discrete alarms
   1: 'Rockwell PLC Comm Fault', class No Acknowledgement, trigger "DB302_HMI_Faults_SDC_Faults_0" bit 0
   2: 'Wireless Access Point 1 Comm Fault', class No Acknowledgement, trigger "DB302_HMI_Faults_SDC_Faults_0" bit 1
   3: 'Wireless Access Point 2 Comm Fault', class No Acknowledgement, trigger "DB302_HMI_Faults_SDC_Faults_0" bit 2
   5: 'Wireless Access Point 4 Comm Fault', class No Acknowledgement, trigger "DB302_HMI_Faults_SDC_Faults_0" bit 4
   6: 'Wireless Access Point 5 Comm Fault', class No Acknowledgement, trigger "DB302_HMI_Faults_SDC_Faults_0" bit 5
   7: 'Wireless Access Point 6 Comm Fault', class No Acknowledgement, trigger "DB302_HMI_Faults_SDC_Faults_0" bit 6
   8: 'Wireless Access Point 7 Comm Fault', class No Acknowledgement, trigger "DB302_HMI_Faults_SDC_Faults_0" bit 7
   9: 'Wireless Access Point 8 Comm Fault', class No Acknowledgement, trigger "DB302_HMI_Faults_SDC_Faults_0" bit 8
   10: 'Wireless Access Point 9 Comm Fault', class No Acknowledgement, trigger "DB302_HMI_Faults_SDC_Faults_0" bit 9
   11: 'Wireless Access Point 10 Comm Fault', class No Acknowledgement, trigger "DB302_HMI_Faults_SDC_Faults_0" bit 10
   12: 'Wireless Access Point 11 Comm Fault', class No Acknowledgement, trigger "DB302_HMI_Faults_SDC_Faults_0" bit 11
   13: 'Wireless Access Point 12 Comm Fault', class No Acknowledgement, trigger "DB302_HMI_Faults_SDC_Faults_0" bit 12
   14: 'Wireless Access Point 13 Comm Fault', class No Acknowledgement, trigger "DB302_HMI_Faults_SDC_Faults_0" bit 13
   15: 'Wireless Access Point 14 Comm Fault', class No Acknowledgement, trigger "DB302_HMI_Faults_SDC_Faults_0" bit 14
   16: 'Wireless Access Point 15 Comm Fault', class No Acknowledgement, trigger "DB302_HMI_Faults_SDC_Faults_0" bit 15
   17: 'Wireless Access Point 16 Comm Fault', class No Acknowledgement, trigger "DB302_HMI_Faults_SDC_Faults_1" bit 0
   18: 'Wireless Access Point 17 Comm Fault', class No Acknowledgement, trigger "DB302_HMI_Faults_SDC_Faults_1" bit 1
   19: 'Wireless Access Point 18 Comm Fault', class No Acknowledgement, trigger "DB302_HMI_Faults_SDC_Faults_1" bit 2
   20: 'Wireless Access Point 19 Comm Fault', class No Acknowledgement, trigger "DB302_HMI_Faults_SDC_Faults_1" bit 3
   21: 'Spare_Fault_021', class No Acknowledgement, trigger "DB302_HMI_Faults_SDC_Faults_1" bit 4
   22: 'Spare_Fault_022', class No Acknowledgement, trigger "DB302_HMI_Faults_SDC_Faults_1" bit 5
   23: 'Spare_Fault_023', class No Acknowledgement, trigger "DB302_HMI_Faults_SDC_Faults_1" bit 6
   24: 'Spare_Fault_024', class No Acknowledgement, trigger "DB302_HMI_Faults_SDC_Faults_1" bit 7
   25: 'Duplicate Carrier Fault', class No Acknowledgement, trigger "DB302_HMI_Faults_SDC_Faults_1" bit 8
   26: 'Spare_Fault_026', class No Acknowledgement, trigger "DB302_HMI_Faults_SDC_Faults_1" bit 9
   27: 'EMS01 System E-Stop', class No Acknowledgement, trigger "DB302_HMI_Faults_SDC_Faults_1" bit 10
   28: 'Spare_Fault_028', class No Acknowledgement, trigger "DB302_HMI_Faults_SDC_Faults_1" bit 11
   29: 'Spare_Fault_029', class No Acknowledgement, trigger "DB302_HMI_Faults_SDC_Faults_1" bit 12
   30: 'Spare_Fault_030', class No Acknowledgement, trigger "DB302_HMI_Faults_SDC_Faults_1" bit 13
   31: 'Spare_Fault_031', class No Acknowledgement, trigger "DB302_HMI_Faults_SDC_Faults_1" bit 14
   32: 'Spare_Fault_032', class No Acknowledgement, trigger "DB302_HMI_Faults_SDC_Faults_1" bit 15
   33: 'Spare_Fault_033', class No Acknowledgement, trigger "DB302_HMI_Faults_SDC_Faults_2" bit 0
   34: 'Spare_Fault_034', class No Acknowledgement, trigger "DB302_HMI_Faults_SDC_Faults_2" bit 1
   35: 'Spare_Fault_035', class No Acknowledgement, trigger "DB302_HMI_Faults_SDC_Faults_2" bit 2
   36: 'Spare_Fault_036', class No Acknowledgement, trigger "DB302_HMI_Faults_SDC_Faults_2" bit 3
   37: 'Spare_Fault_037', class No Acknowledgement, trigger "DB302_HMI_Faults_SDC_Faults_2" bit 4
   38: 'Spare_Fault_038', class No Acknowledgement, trigger "DB302_HMI_Faults_SDC_Faults_2" bit 5
   39: 'Spare_Fault_039', class No Acknowledgement, trigger "DB302_HMI_Faults_SDC_Faults_2" bit 6
   40: 'Spare_Fault_040', class No Acknowledgement, trigger "DB302_HMI_Faults_SDC_Faults_2" bit 7
   41: 'Spare_Fault_041', class No Acknowledgement, trigger "DB302_HMI_Faults_SDC_Faults_2" bit 8
   42: 'Spare_Fault_042', class No Acknowledgement, trigger "DB302_HMI_Faults_SDC_Faults_2" bit 9
   43: 'Spare_Fault_043', class No Acknowledgement, trigger "DB302_HMI_Faults_SDC_Faults_2" bit 10
   44: 'Spare_Fault_044', class No Acknowledgement, trigger "DB302_HMI_Faults_SDC_Faults_2" bit 11
   45: 'Spare_Fault_045', class No Acknowledgement, trigger "DB302_HMI_Faults_SDC_Faults_2" bit 12
   46: 'Spare_Fault_046', class No Acknowledgement, trigger "DB302_HMI_Faults_SDC_Faults_2" bit 13
   47: 'Spare_Fault_047', class No Acknowledgement, trigger "DB302_HMI_Faults_SDC_Faults_2" bit 14
   48: 'Spare_Fault_048', class No Acknowledgement, trigger "DB302_HMI_Faults_SDC_Faults_2" bit 15
   49: 'Spare_Fault_049', class No Acknowledgement, trigger "DB302_HMI_Faults_SDC_Faults_3" bit 0
   50: 'Spare_Fault_050', class No Acknowledgement, trigger "DB302_HMI_Faults_SDC_Faults_3" bit 1
   51: 'Spare_Fault_051', class No Acknowledgement, trigger "DB302_HMI_Faults_SDC_Faults_3" bit 2
   52: 'Spare_Fault_052', class No Acknowledgement, trigger "DB302_HMI_Faults_SDC_Faults_3" bit 3
   53: 'Spare_Fault_053', class No Acknowledgement, trigger "DB302_HMI_Faults_SDC_Faults_3" bit 4
   54: 'Spare_Fault_054', class No Acknowledgement, trigger "DB302_HMI_Faults_SDC_Faults_3" bit 5
   55: 'Spare_Fault_055', class No Acknowledgement, trigger "DB302_HMI_Faults_SDC_Faults_3" bit 6
   56: 'Spare_Fault_056', class No Acknowledgement, trigger "DB302_HMI_Faults_SDC_Faults_3" bit 7
   57: 'Spare_Fault_057', class No Acknowledgement, trigger "DB302_HMI_Faults_SDC_Faults_3" bit 8
   58: 'Spare_Fault_058', class No Acknowledgement, trigger "DB302_HMI_Faults_SDC_Faults_3" bit 9
   59: 'Spare_Fault_059', class No Acknowledgement, trigger "DB302_HMI_Faults_SDC_Faults_3" bit 10
   60: 'Spare_Fault_060', class No Acknowledgement, trigger "DB302_HMI_Faults_SDC_Faults_3" bit 11
   61: 'Spare_Fault_061', class No Acknowledgement, trigger "DB302_HMI_Faults_SDC_Faults_3" bit 12
   62: 'Spare_Fault_062', class No Acknowledgement, trigger "DB302_HMI_Faults_SDC_Faults_3" bit 13
   63: 'Spare_Fault_063', class No Acknowledgement, trigger "DB302_HMI_Faults_SDC_Faults_3" bit 14
   64: 'Spare_Fault_064', class No Acknowledgement, trigger "DB302_HMI_Faults_SDC_Faults_3" bit 15
   65: 'Carrier 01 Disconnect Open Power Fault DI11.0', class No Acknowledgement, trigger "DB302_HMI_Faults_Carrier1_Faults_0" bit 0
   66: 'Carrier 01 Drive Profinet Comm Fault', class No Acknowledgement, trigger "DB302_HMI_Faults_Carrier1_Faults_0" bit 1
   67: 'Carrier 01 Production Stop Not Reset', class No Acknowledgement, trigger "DB302_HMI_Faults_Carrier1_Faults_0" bit 2
   68: 'Carrier 01 CB02122 Tripped', class No Acknowledgement, trigger "DB302_HMI_Faults_Carrier1_Faults_0" bit 3
   69: 'Carrier 01 CB02123 Tripped', class No Acknowledgement, trigger "DB302_HMI_Faults_Carrier1_Faults_0" bit 4
   70: 'Carrier 01 AUX1 CB Tripped', class No Acknowledgement, trigger "DB302_HMI_Faults_Carrier1_Faults_0" bit 5
   71: 'Carrier 01 AUX2 CB Tripped', class No Acknowledgement, trigger "DB302_HMI_Faults_Carrier1_Faults_0" bit 6
   72: 'Carrier 01 PLC Not Communicating', class No Acknowledgement, trigger "DB302_HMI_Faults_Carrier1_Faults_0" bit 7
   73: 'Carrier 01 Safe Input Card Fault', class No Acknowledgement, trigger "DB302_HMI_Faults_Carrier1_Faults_0" bit 8
   74: 'Carrier 01 Safe Output Card Fault', class No Acknowledgement, trigger "DB302_HMI_Faults_Carrier1_Faults_0" bit 9
   75: 'Carrier 01 Standard Input Card Fault', class No Acknowledgement, trigger "DB302_HMI_Faults_Carrier1_Faults_0" bit 10
   76: 'Carrier 01 Standard Output Card Fault', class No Acknowledgement, trigger "DB302_HMI_Faults_Carrier1_Faults_0" bit 11
   77: 'Carrier 01 Encoder Position Fault', class No Acknowledgement, trigger "DB302_HMI_Faults_Carrier1_Faults_0" bit 12
   78: 'Carrier 01 Encoder Internal Error', class No Acknowledgement, trigger "DB302_HMI_Faults_Carrier1_Faults_0" bit 13
   79: 'Carrier 01 Encoder Comm Fault', class No Acknowledgement, trigger "DB302_HMI_Faults_Carrier1_Faults_0" bit 14
   80: 'Carrier 01 HMI Comm Fault', class No Acknowledgement, trigger "DB302_HMI_Faults_Carrier1_Faults_0" bit 15
   81: 'Carrier 01 Crash Detection Fault', class No Acknowledgement, trigger "DB302_HMI_Faults_Carrier1_Faults_1" bit 0
   82: 'Carrier 01 Carrier Number Invalid', class No Acknowledgement, trigger "DB302_HMI_Faults_Carrier1_Faults_1" bit 1
   83: 'Carrier 01 Drive: PROFINET configuration error', class No Acknowledgement, trigger "DB302_HMI_Faults_Carrier1_Faults_1" bit 2
   84: 'Carrier 01 Drive: Error internal communications', class No Acknowledgement, trigger "DB302_HMI_Faults_Carrier1_Faults_1" bit 3
   85: 'Carrier 01 Drive: Motor overtemperature', class No Acknowledgement, trigger "DB302_HMI_Faults_Carrier1_Faults_1" bit 4
   86: 'Carrier 01 Drive: Motor overcurrent', class No Acknowledgement, trigger "DB302_HMI_Faults_Carrier1_Faults_1" bit 5
   87: 'Carrier 01 Drive: Infeed or power unit not ready', class No Acknowledgement, trigger "DB302_HMI_Faults_Carrier1_Faults_1" bit 6
   88: 'Carrier 01 Drive: Short-circuit/ground fault detected', class No Acknowledgement, trigger "DB302_HMI_Faults_Carrier1_Faults_1" bit 7
   89: 'Carrier 01 Drive: PROFINET Setpoint timeout', class No Acknowledgement, trigger "DB302_HMI_Faults_Carrier1_Faults_1" bit 8
   90: 'Carrier 01 Power unit: Overcurrent', class No Acknowledgement, trigger "DB302_HMI_Faults_Carrier1_Faults_1" bit 9
   91: 'Carrier 01 Power unit: DC link voltage overvoltage', class No Acknowledgement, trigger "DB302_HMI_Faults_Carrier1_Faults_1" bit 10
   92: 'Carrier 01 Power unit: DC link voltage undervoltage', class No Acknowledgement, trigger "DB302_HMI_Faults_Carrier1_Faults_1" bit 11
   93: 'Carrier 01 Power unit: Line phase failure in main circuit', class No Acknowledgement, trigger "DB302_HMI_Faults_Carrier1_Faults_1" bit 12
   94: 'Carrier 01 Power unit: Phase failure motor cable', class No Acknowledgement, trigger "DB302_HMI_Faults_Carrier1_Faults_1" bit 13
   95: 'Carrier 01 Power unit: Ground fault', class No Acknowledgement, trigger "DB302_HMI_Faults_Carrier1_Faults_1" bit 14
   96: 'Spare_Fault_096', class No Acknowledgement, trigger "DB302_HMI_Faults_Carrier1_Faults_1" bit 15
   97: 'Carrier 01 Motion Off Fault', class No Acknowledgement, trigger "DB302_HMI_Faults_Carrier1_Faults_2" bit 0
   98: 'Carrier 01 Motion On Fault', class No Acknowledgement, trigger "DB302_HMI_Faults_Carrier1_Faults_2" bit 1
   99: 'Carrier 01 Spacing Fault', class No Acknowledgement, trigger "DB302_HMI_Faults_Carrier1_Faults_2" bit 2
   100: 'Carrier 01 Duplicate Carrier Number Fault', class No Acknowledgement, trigger "DB302_HMI_Faults_Carrier1_Faults_2" bit 3
   101: 'Spare_Fault_101', class No Acknowledgement, trigger "DB302_HMI_Faults_Carrier1_Faults_2" bit 4
   102: 'Spare_Fault_102', class No Acknowledgement, trigger "DB302_HMI_Faults_Carrier1_Faults_2" bit 5
   103: 'Spare_Fault_103', class No Acknowledgement, trigger "DB302_HMI_Faults_Carrier1_Faults_2" bit 6
   104: 'Spare_Fault_104', class No Acknowledgement, trigger "DB302_HMI_Faults_Carrier1_Faults_2" bit 7
   105: 'Spare_Fault_105', class No Acknowledgement, trigger "DB302_HMI_Faults_Carrier1_Faults_2" bit 8
   106: 'Spare_Fault_106', class No Acknowledgement, trigger "DB302_HMI_Faults_Carrier1_Faults_2" bit 9
   107: 'Spare_Fault_107', class No Acknowledgement, trigger "DB302_HMI_Faults_Carrier1_Faults_2" bit 10
   108: 'Spare_Fault_108', class No Acknowledgement, trigger "DB302_HMI_Faults_Carrier1_Faults_2" bit 11
   109: 'Spare_Fault_109', class No Acknowledgement, trigger "DB302_HMI_Faults_Carrier1_Faults_2" bit 12
   110: 'Spare_Fault_110', class No Acknowledgement, trigger "DB302_HMI_Faults_Carrier1_Faults_2" bit 13
   111: 'Spare_Fault_111', class No Acknowledgement, trigger "DB302_HMI_Faults_Carrier1_Faults_2" bit 14
   112: 'Spare_Fault_112', class No Acknowledgement, trigger "DB302_HMI_Faults_Carrier1_Faults_2" bit 15
   113: 'Spare_Fault_113', class No Acknowledgement, trigger "DB302_HMI_Faults_Carrier1_Faults_3" bit 0
   114: 'Spare_Fault_114', class No Acknowledgement, trigger "DB302_HMI_Faults_Carrier1_Faults_3" bit 1
   115: 'Spare_Fault_115', class No Acknowledgement, trigger "DB302_HMI_Faults_Carrier1_Faults_3" bit 2
   116: 'Spare_Fault_116', class No Acknowledgement, trigger "DB302_HMI_Faults_Carrier1_Faults_3" bit 3
   117: 'Spare_Fault_117', class No Acknowledgement, trigger "DB302_HMI_Faults_Carrier1_Faults_3" bit 4
   118: 'Spare_Fault_118', class No Acknowledgement, trigger "DB302_HMI_Faults_Carrier1_Faults_3" bit 5
   119: 'Spare_Fault_119', class No Acknowledgement, trigger "DB302_HMI_Faults_Carrier1_Faults_3" bit 6
   120: 'Spare_Fault_120', class No Acknowledgement, trigger "DB302_HMI_Faults_Carrier1_Faults_3" bit 7
   121: 'Spare_Fault_121', class No Acknowledgement, trigger "DB302_HMI_Faults_Carrier1_Faults_3" bit 8
   122: 'Spare_Fault_122', class No Acknowledgement, trigger "DB302_HMI_Faults_Carrier1_Faults_3" bit 9
   123: 'Spare_Fault_123', class No Acknowledgement, trigger "DB302_HMI_Faults_Carrier1_Faults_3" bit 10
   124: 'Spare_Fault_124', class No Acknowledgement, trigger "DB302_HMI_Faults_Carrier1_Faults_3" bit 11
   125: 'Spare_Fault_125', class No Acknowledgement, trigger "DB302_HMI_Faults_Carrier1_Faults_3" bit 12
   126: 'Spare_Fault_126', class No Acknowledgement, trigger "DB302_HMI_Faults_Carrier1_Faults_3" bit 13
   127: 'Spare_Fault_127', class No Acknowledgement, trigger "DB302_HMI_Faults_Carrier1_Faults_3" bit 14
   128: 'Spare_Fault_128', class No Acknowledgement, trigger "DB302_HMI_Faults_Carrier1_Faults_3" bit 15
   129: 'Carrier 02 Disconnect Open Power Fault DI11.0', class No Acknowledgement, trigger "DB302_HMI_Faults_Carrier2_Faults_0" bit 0
   130: 'Carrier 02 Drive Profinet Comm Fault', class No Acknowledgement, trigger "DB302_HMI_Faults_Carrier2_Faults_0" bit 1
   131: 'Carrier 02 Production Stop Not Reset', class No Acknowledgement, trigger "DB302_HMI_Faults_Carrier2_Faults_0" bit 2
   132: 'Carrier 02 CB02122 Tripped', class No Acknowledgement, trigger "DB302_HMI_Faults_Carrier2_Faults_0" bit 3
   133: 'Carrier 02 CB02123 Tripped', class No Acknowledgement, trigger "DB302_HMI_Faults_Carrier2_Faults_0" bit 4
   134: 'Carrier 02 AUX1 CB Tripped', class No Acknowledgement, trigger "DB302_HMI_Faults_Carrier2_Faults_0" bit 5
   135: 'Carrier 02 AUX2 CB Tripped', class No Acknowledgement, trigger "DB302_HMI_Faults_Carrier2_Faults_0" bit 6
   136: 'Carrier 02 PLC Not Communicating', class No Acknowledgement, trigger "DB302_HMI_Faults_Carrier2_Faults_0" bit 7
   137: 'Carrier 02 Safe Input Card Fault', class No Acknowledgement, trigger "DB302_HMI_Faults_Carrier2_Faults_0" bit 8
   138: 'Carrier 02 Safe Output Card Fault', class No Acknowledgement, trigger "DB302_HMI_Faults_Carrier2_Faults_0" bit 9
   139: 'Carrier 02 Standard Input Card Fault', class No Acknowledgement, trigger "DB302_HMI_Faults_Carrier2_Faults_0" bit 10
   140: 'Carrier 02 Standard Output Card Fault', class No Acknowledgement, trigger "DB302_HMI_Faults_Carrier2_Faults_0" bit 11
   141: 'Carrier 02 Encoder Position Fault', class No Acknowledgement, trigger "DB302_HMI_Faults_Carrier2_Faults_0" bit 12
   142: 'Carrier 02 Encoder Internal Error', class No Acknowledgement, trigger "DB302_HMI_Faults_Carrier2_Faults_0" bit 13
   143: 'Carrier 02 Encoder Comm Fault', class No Acknowledgement, trigger "DB302_HMI_Faults_Carrier2_Faults_0" bit 14
   144: 'Carrier 02 HMI Comm Fault', class No Acknowledgement, trigger "DB302_HMI_Faults_Carrier2_Faults_0" bit 15
   145: 'Carrier 02 Crash Detection Fault', class No Acknowledgement, trigger "DB302_HMI_Faults_Carrier2_Faults_1" bit 0
   146: 'Carrier 02 Carrier Number Invalid', class No Acknowledgement, trigger "DB302_HMI_Faults_Carrier2_Faults_1" bit 1
   147: 'Carrier 02 Drive: PROFINET configuration error', class No Acknowledgement, trigger "DB302_HMI_Faults_Carrier2_Faults_1" bit 2
   148: 'Carrier 02 Drive: Error internal communications', class No Acknowledgement, trigger "DB302_HMI_Faults_Carrier2_Faults_1" bit 3
   149: 'Carrier 02 Drive: Motor overtemperature', class No Acknowledgement, trigger "DB302_HMI_Faults_Carrier2_Faults_1" bit 4
   150: 'Carrier 02 Drive: Motor overcurrent', class No Acknowledgement, trigger "DB302_HMI_Faults_Carrier2_Faults_1" bit 5
   151: 'Carrier 02 Drive: Infeed or power unit not ready', class No Acknowledgement, trigger "DB302_HMI_Faults_Carrier2_Faults_1" bit 6
   152: 'Carrier 02 Drive: Short-circuit/ground fault detected', class No Acknowledgement, trigger "DB302_HMI_Faults_Carrier2_Faults_1" bit 7
   153: 'Carrier 02 Drive: PROFINET Setpoint timeout', class No Acknowledgement, trigger "DB302_HMI_Faults_Carrier2_Faults_1" bit 8
   154: 'Carrier 02 Power unit: Overcurrent', class No Acknowledgement, trigger "DB302_HMI_Faults_Carrier2_Faults_1" bit 9
   155: 'Carrier 02 Power unit: DC link voltage overvoltage', class No Acknowledgement, trigger "DB302_HMI_Faults_Carrier2_Faults_1" bit 10
   156: 'Carrier 02 Power unit: DC link voltage undervoltage', class No Acknowledgement, trigger "DB302_HMI_Faults_Carrier2_Faults_1" bit 11
   157: 'Carrier 02 Power unit: Line phase failure in main circuit', class No Acknowledgement, trigger "DB302_HMI_Faults_Carrier2_Faults_1" bit 12
   158: 'Carrier 02 Power unit: Phase failure motor cable', class No Acknowledgement, trigger "DB302_HMI_Faults_Carrier2_Faults_1" bit 13
   159: 'Carrier 02 Power unit: Ground fault', class No Acknowledgement, trigger "DB302_HMI_Faults_Carrier2_Faults_1" bit 14
   160: 'Spare_Fault_160', class No Acknowledgement, trigger "DB302_HMI_Faults_Carrier2_Faults_1" bit 15
   161: 'Carrier 02 Motion Off Fault', class No Acknowledgement, trigger "DB302_HMI_Faults_Carrier2_Faults_2" bit 0
   162: 'Carrier 02 Motion On Fault', class No Acknowledgement, trigger "DB302_HMI_Faults_Carrier2_Faults_2" bit 1
   163: 'Carrier 02 Spacing Fault', class No Acknowledgement, trigger "DB302_HMI_Faults_Carrier2_Faults_2" bit 2
   164: 'Carrier 02 Duplicate Carrier Number Fault', class No Acknowledgement, trigger "DB302_HMI_Faults_Carrier2_Faults_2" bit 3
   165: 'Spare_Fault_165', class No Acknowledgement, trigger "DB302_HMI_Faults_Carrier2_Faults_2" bit 4
   166: 'Spare_Fault_166', class No Acknowledgement, trigger "DB302_HMI_Faults_Carrier2_Faults_2" bit 5
   167: 'Spare_Fault_167', class No Acknowledgement, trigger "DB302_HMI_Faults_Carrier2_Faults_2" bit 6
   168: 'Spare_Fault_168', class No Acknowledgement, trigger "DB302_HMI_Faults_Carrier2_Faults_2" bit 7
   169: 'Spare_Fault_169', class No Acknowledgement, trigger "DB302_HMI_Faults_Carrier2_Faults_2" bit 8
   170: 'Spare_Fault_170', class No Acknowledgement, trigger "DB302_HMI_Faults_Carrier2_Faults_2" bit 9
   171: 'Spare_Fault_171', class No Acknowledgement, trigger "DB302_HMI_Faults_Carrier2_Faults_2" bit 10
   172: 'Spare_Fault_172', class No Acknowledgement, trigger "DB302_HMI_Faults_Carrier2_Faults_2" bit 11
   173: 'Spare_Fault_173', class No Acknowledgement, trigger "DB302_HMI_Faults_Carrier2_Faults_2" bit 12
   174: 'Spare_Fault_174', class No Acknowledgement, trigger "DB302_HMI_Faults_Carrier2_Faults_2" bit 13
   175: 'Spare_Fault_175', class No Acknowledgement, trigger "DB302_HMI_Faults_Carrier2_Faults_2" bit 14
   176: 'Spare_Fault_176', class No Acknowledgement, trigger "DB302_HMI_Faults_Carrier2_Faults_2" bit 15
   177: 'Spare_Fault_177', class No Acknowledgement, trigger "DB302_HMI_Faults_Carrier2_Faults_3" bit 0
   178: 'Spare_Fault_178', class No Acknowledgement, trigger "DB302_HMI_Faults_Carrier2_Faults_3" bit 1
   179: 'Spare_Fault_179', class No Acknowledgement, trigger "DB302_HMI_Faults_Carrier2_Faults_3" bit 2
   180: 'Spare_Fault_180', class No Acknowledgement, trigger "DB302_HMI_Faults_Carrier2_Faults_3" bit 3
   181: 'Spare_Fault_181', class No Acknowledgement, trigger "DB302_HMI_Faults_Carrier2_Faults_3" bit 4
   182: 'Spare_Fault_182', class No Acknowledgement, trigger "DB302_HMI_Faults_Carrier2_Faults_3" bit 5
   183: 'Spare_Fault_183', class No Acknowledgement, trigger "DB302_HMI_Faults_Carrier2_Faults_3" bit 6
   184: 'Spare_Fault_184', class No Acknowledgement, trigger "DB302_HMI_Faults_Carrier2_Faults_3" bit 7
   185: 'Spare_Fault_185', class No Acknowledgement, trigger "DB302_HMI_Faults_Carrier2_Faults_3" bit 8
   186: 'Spare_Fault_186', class No Acknowledgement, trigger "DB302_HMI_Faults_Carrier2_Faults_3" bit 9
   187: 'Spare_Fault_187', class No Acknowledgement, trigger "DB302_HMI_Faults_Carrier2_Faults_3" bit 10
   188: 'Spare_Fault_188', class No Acknowledgement, trigger "DB302_HMI_Faults_Carrier2_Faults_3" bit 11
   189: 'Spare_Fault_189', class No Acknowledgement, trigger "DB302_HMI_Faults_Carrier2_Faults_3" bit 12
   190: 'Spare_Fault_190', class No Acknowledgement, trigger "DB302_HMI_Faults_Carrier2_Faults_3" bit 13
   191: 'Spare_Fault_191', class No Acknowledgement, trigger "DB302_HMI_Faults_Carrier2_Faults_3" bit 14
   192: 'Spare_Fault_192', class No Acknowledgement, trigger "DB302_HMI_Faults_Carrier2_Faults_3" bit 15
   193: 'Carrier 03 Disconnect Open Power Fault DI11.0', class No Acknowledgement, trigger "DB302_HMI_Faults_Carrier3_Faults_0" bit 0
   194: 'Carrier 03 Drive Profinet Comm Fault', class No Acknowledgement, trigger "DB302_HMI_Faults_Carrier3_Faults_0" bit 1
   195: 'Carrier 03 Production Stop Not Reset', class No Acknowledgement, trigger "DB302_HMI_Faults_Carrier3_Faults_0" bit 2
   196: 'Carrier 03 CB02122 Tripped', class No Acknowledgement, trigger "DB302_HMI_Faults_Carrier3_Faults_0" bit 3
   197: 'Carrier 03 CB02123 Tripped', class No Acknowledgement, trigger "DB302_HMI_Faults_Carrier3_Faults_0" bit 4
   198: 'Carrier 03 AUX1 CB Tripped', class No Acknowledgement, trigger "DB302_HMI_Faults_Carrier3_Faults_0" bit 5
   199: 'Carrier 03 AUX2 CB Tripped', class No Acknowledgement, trigger "DB302_HMI_Faults_Carrier3_Faults_0" bit 6
   200: 'Carrier 03 PLC Not Communicating', class No Acknowledgement, trigger "DB302_HMI_Faults_Carrier3_Faults_0" bit 7
   201: 'Carrier 03 Safe Input Card Fault', class No Acknowledgement, trigger "DB302_HMI_Faults_Carrier3_Faults_0" bit 8
   202: 'Carrier 03 Safe Output Card Fault', class No Acknowledgement, trigger "DB302_HMI_Faults_Carrier3_Faults_0" bit 9
   203: 'Carrier 03 Standard Input Card Fault', class No Acknowledgement, trigger "DB302_HMI_Faults_Carrier3_Faults_0" bit 10
   204: 'Carrier 03 Standard Output Card Fault', class No Acknowledgement, trigger "DB302_HMI_Faults_Carrier3_Faults_0" bit 11
   205: 'Carrier 03 Encoder Position Fault', class No Acknowledgement, trigger "DB302_HMI_Faults_Carrier3_Faults_0" bit 12
   206: 'Carrier 03 Encoder Internal Error', class No Acknowledgement, trigger "DB302_HMI_Faults_Carrier3_Faults_0" bit 13
   207: 'Carrier 03 Encoder Comm Fault', class No Acknowledgement, trigger "DB302_HMI_Faults_Carrier3_Faults_0" bit 14
   208: 'Carrier 03 HMI Comm Fault', class No Acknowledgement, trigger "DB302_HMI_Faults_Carrier3_Faults_0" bit 15
   209: 'Carrier 03 Crash Detection Fault', class No Acknowledgement, trigger "DB302_HMI_Faults_Carrier3_Faults_1" bit 0
   210: 'Carrier 03 Carrier Number Invalid', class No Acknowledgement, trigger "DB302_HMI_Faults_Carrier3_Faults_1" bit 1
   211: 'Carrier 03 Drive: PROFINET configuration error', class No Acknowledgement, trigger "DB302_HMI_Faults_Carrier3_Faults_1" bit 2
   212: 'Carrier 03 Drive: Error internal communications', class No Acknowledgement, trigger "DB302_HMI_Faults_Carrier3_Faults_1" bit 3
   213: 'Carrier 03 Drive: Motor overtemperature', class No Acknowledgement, trigger "DB302_HMI_Faults_Carrier3_Faults_1" bit 4
   214: 'Carrier 03 Drive: Motor overcurrent', class No Acknowledgement, trigger "DB302_HMI_Faults_Carrier3_Faults_1" bit 5
   215: 'Carrier 03 Drive: Infeed or power unit not ready', class No Acknowledgement, trigger "DB302_HMI_Faults_Carrier3_Faults_1" bit 6
   216: 'Carrier 03 Drive: Short-circuit/ground fault detected', class No Acknowledgement, trigger "DB302_HMI_Faults_Carrier3_Faults_1" bit 7
   217: 'Carrier 03 Drive: PROFINET Setpoint timeout', class No Acknowledgement, trigger "DB302_HMI_Faults_Carrier3_Faults_1" bit 8
   218: 'Carrier 03 Power unit: Overcurrent', class No Acknowledgement, trigger "DB302_HMI_Faults_Carrier3_Faults_1" bit 9
   219: 'Carrier 03 Power unit: DC link voltage overvoltage', class No Acknowledgement, trigger "DB302_HMI_Faults_Carrier3_Faults_1" bit 10
   220: 'Carrier 03 Power unit: DC link voltage undervoltage', class No Acknowledgement, trigger "DB302_HMI_Faults_Carrier3_Faults_1" bit 11
   221: 'Carrier 03 Power unit: Line phase failure in main circuit', class No Acknowledgement, trigger "DB302_HMI_Faults_Carrier3_Faults_1" bit 12
   222: 'Carrier 03 Power unit: Phase failure motor cable', class No Acknowledgement, trigger "DB302_HMI_Faults_Carrier3_Faults_1" bit 13
   223: 'Carrier 03 Power unit: Ground fault', class No Acknowledgement, trigger "DB302_HMI_Faults_Carrier3_Faults_1" bit 14
   224: 'Spare_Fault_224', class No Acknowledgement, trigger "DB302_HMI_Faults_Carrier3_Faults_1" bit 15
   225: 'Carrier 03 Motion Off Fault', class No Acknowledgement, trigger "DB302_HMI_Faults_Carrier3_Faults_2" bit 0
   226: 'Carrier 03 Motion On Fault', class No Acknowledgement, trigger "DB302_HMI_Faults_Carrier3_Faults_2" bit 1
   227: 'Carrier 03 Spacing Fault', class No Acknowledgement, trigger "DB302_HMI_Faults_Carrier3_Faults_2" bit 2
   228: 'Carrier 03 Duplicate Carrier Number Fault', class No Acknowledgement, trigger "DB302_HMI_Faults_Carrier3_Faults_2" bit 3
   229: 'Spare_Fault_229', class No Acknowledgement, trigger "DB302_HMI_Faults_Carrier3_Faults_2" bit 4
   230: 'Spare_Fault_230', class No Acknowledgement, trigger "DB302_HMI_Faults_Carrier3_Faults_2" bit 5
   231: 'Spare_Fault_231', class No Acknowledgement, trigger "DB302_HMI_Faults_Carrier3_Faults_2" bit 6
   232: 'Spare_Fault_232', class No Acknowledgement, trigger "DB302_HMI_Faults_Carrier3_Faults_2" bit 7
   233: 'Spare_Fault_233', class No Acknowledgement, trigger "DB302_HMI_Faults_Carrier3_Faults_2" bit 8
   234: 'Spare_Fault_234', class No Acknowledgement, trigger "DB302_HMI_Faults_Carrier3_Faults_2" bit 9
   235: 'Spare_Fault_235', class No Acknowledgement, trigger "DB302_HMI_Faults_Carrier3_Faults_2" bit 10
   236: 'Spare_Fault_236', class No Acknowledgement, trigger "DB302_HMI_Faults_Carrier3_Faults_2" bit 11
   237: 'Spare_Fault_237', class No Acknowledgement, trigger "DB302_HMI_Faults_Carrier3_Faults_2" bit 12
   238: 'Spare_Fault_238', class No Acknowledgement, trigger "DB302_HMI_Faults_Carrier3_Faults_2" bit 13
   239: 'Spare_Fault_239', class No Acknowledgement, trigger "DB302_HMI_Faults_Carrier3_Faults_2" bit 14
   240: 'Spare_Fault_240', class No Acknowledgement, trigger "DB302_HMI_Faults_Carrier3_Faults_2" bit 15
   241: 'Spare_Fault_241', class No Acknowledgement, trigger "DB302_HMI_Faults_Carrier3_Faults_3" bit 0
   242: 'Spare_Fault_242', class No Acknowledgement, trigger "DB302_HMI_Faults_Carrier3_Faults_3" bit 1
   243: 'Spare_Fault_243', class No Acknowledgement, trigger "DB302_HMI_Faults_Carrier3_Faults_3" bit 2
   244: 'Spare_Fault_244', class No Acknowledgement, trigger "DB302_HMI_Faults_Carrier3_Faults_3" bit 3
   245: 'Spare_Fault_245', class No Acknowledgement, trigger "DB302_HMI_Faults_Carrier3_Faults_3" bit 4
   246: 'Spare_Fault_246', class No Acknowledgement, trigger "DB302_HMI_Faults_Carrier3_Faults_3" bit 5
   247: 'Spare_Fault_247', class No Acknowledgement, trigger "DB302_HMI_Faults_Carrier3_Faults_3" bit 6
   248: 'Spare_Fault_248', class No Acknowledgement, trigger "DB302_HMI_Faults_Carrier3_Faults_3" bit 7
   249: 'Spare_Fault_249', class No Acknowledgement, trigger "DB302_HMI_Faults_Carrier3_Faults_3" bit 8
   250: 'Spare_Fault_250', class No Acknowledgement, trigger "DB302_HMI_Faults_Carrier3_Faults_3" bit 9
   251: 'Spare_Fault_251', class No Acknowledgement, trigger "DB302_HMI_Faults_Carrier3_Faults_3" bit 10
   252: 'Spare_Fault_252', class No Acknowledgement, trigger "DB302_HMI_Faults_Carrier3_Faults_3" bit 11
   253: 'Spare_Fault_253', class No Acknowledgement, trigger "DB302_HMI_Faults_Carrier3_Faults_3" bit 12
   254: 'Spare_Fault_254', class No Acknowledgement, trigger "DB302_HMI_Faults_Carrier3_Faults_3" bit 13
   255: 'Spare_Fault_255', class No Acknowledgement, trigger "DB302_HMI_Faults_Carrier3_Faults_3" bit 14
   256: 'Spare_Fault_256', class No Acknowledgement, trigger "DB302_HMI_Faults_Carrier3_Faults_3" bit 15
   257: 'Carrier 04 Disconnect Open Power Fault DI11.0', class No Acknowledgement, trigger "DB302_HMI_Faults_Carrier4_Faults_0" bit 0
   258: 'Carrier 04 Drive Profinet Comm Fault', class No Acknowledgement, trigger "DB302_HMI_Faults_Carrier4_Faults_0" bit 1
   259: 'Carrier 04 Production Stop Not Reset', class No Acknowledgement, trigger "DB302_HMI_Faults_Carrier4_Faults_0" bit 2
   260: 'Carrier 04 CB02122 Tripped', class No Acknowledgement, trigger "DB302_HMI_Faults_Carrier4_Faults_0" bit 3
   261: 'Carrier 04 CB02123 Tripped', class No Acknowledgement, trigger "DB302_HMI_Faults_Carrier4_Faults_0" bit 4
   262: 'Carrier 04 AUX1 CB Tripped', class No Acknowledgement, trigger "DB302_HMI_Faults_Carrier4_Faults_0" bit 5
   263: 'Carrier 04 AUX2 CB Tripped', class No Acknowledgement, trigger "DB302_HMI_Faults_Carrier4_Faults_0" bit 6
   264: 'Carrier 04 PLC Not Communicating', class No Acknowledgement, trigger "DB302_HMI_Faults_Carrier4_Faults_0" bit 7
   265: 'Carrier 04 Safe Input Card Fault', class No Acknowledgement, trigger "DB302_HMI_Faults_Carrier4_Faults_0" bit 8
   266: 'Carrier 04 Safe Output Card Fault', class No Acknowledgement, trigger "DB302_HMI_Faults_Carrier4_Faults_0" bit 9
   267: 'Carrier 04 Standard Input Card Fault', class No Acknowledgement, trigger "DB302_HMI_Faults_Carrier4_Faults_0" bit 10
   268: 'Carrier 04 Standard Output Card Fault', class No Acknowledgement, trigger "DB302_HMI_Faults_Carrier4_Faults_0" bit 11
   269: 'Carrier 04 Encoder Position Fault', class No Acknowledgement, trigger "DB302_HMI_Faults_Carrier4_Faults_0" bit 12
   270: 'Carrier 04 Encoder Internal Error', class No Acknowledgement, trigger "DB302_HMI_Faults_Carrier4_Faults_0" bit 13
   271: 'Carrier 04 Encoder Comm Fault', class No Acknowledgement, trigger "DB302_HMI_Faults_Carrier4_Faults_0" bit 14
   272: 'Carrier 04 HMI Comm Fault', class No Acknowledgement, trigger "DB302_HMI_Faults_Carrier4_Faults_0" bit 15
   273: 'Carrier 04 Crash Detection Fault', class No Acknowledgement, trigger "DB302_HMI_Faults_Carrier4_Faults_1" bit 0
   274: 'Carrier 04 Carrier Number Invalid', class No Acknowledgement, trigger "DB302_HMI_Faults_Carrier4_Faults_1" bit 1
   275: 'Carrier 04 Drive: PROFINET configuration error', class No Acknowledgement, trigger "DB302_HMI_Faults_Carrier4_Faults_1" bit 2
   276: 'Carrier 04 Drive: Error internal communications', class No Acknowledgement, trigger "DB302_HMI_Faults_Carrier4_Faults_1" bit 3
   277: 'Carrier 04 Drive: Motor overtemperature', class No Acknowledgement, trigger "DB302_HMI_Faults_Carrier4_Faults_1" bit 4
   278: 'Carrier 04 Drive: Motor overcurrent', class No Acknowledgement, trigger "DB302_HMI_Faults_Carrier4_Faults_1" bit 5
   279: 'Carrier 04 Drive: Infeed or power unit not ready', class No Acknowledgement, trigger "DB302_HMI_Faults_Carrier4_Faults_1" bit 6
   280: 'Carrier 04 Drive: Short-circuit/ground fault detected', class No Acknowledgement, trigger "DB302_HMI_Faults_Carrier4_Faults_1" bit 7
   281: 'Carrier 04 Drive: PROFINET Setpoint timeout', class No Acknowledgement, trigger "DB302_HMI_Faults_Carrier4_Faults_1" bit 8
   282: 'Carrier 04 Power unit: Overcurrent', class No Acknowledgement, trigger "DB302_HMI_Faults_Carrier4_Faults_1" bit 9
   283: 'Carrier 04 Power unit: DC link voltage overvoltage', class No Acknowledgement, trigger "DB302_HMI_Faults_Carrier4_Faults_1" bit 10
   284: 'Carrier 04 Power unit: DC link voltage undervoltage', class No Acknowledgement, trigger "DB302_HMI_Faults_Carrier4_Faults_1" bit 11
   285: 'Carrier 04 Power unit: Line phase failure in main circuit', class No Acknowledgement, trigger "DB302_HMI_Faults_Carrier4_Faults_1" bit 12
   286: 'Carrier 04 Power unit: Phase failure motor cable', class No Acknowledgement, trigger "DB302_HMI_Faults_Carrier4_Faults_1" bit 13
   287: 'Carrier 04 Power unit: Ground fault', class No Acknowledgement, trigger "DB302_HMI_Faults_Carrier4_Faults_1" bit 14
   288: 'Spare_Fault_288', class No Acknowledgement, trigger "DB302_HMI_Faults_Carrier4_Faults_1" bit 15
   289: 'Carrier 04 Motion Off Fault', class No Acknowledgement, trigger "DB302_HMI_Faults_Carrier4_Faults_2" bit 0
   290: 'Carrier 04 Motion On Fault', class No Acknowledgement, trigger "DB302_HMI_Faults_Carrier4_Faults_2" bit 1
   291: 'Carrier 04 Spacing Fault', class No Acknowledgement, trigger "DB302_HMI_Faults_Carrier4_Faults_2" bit 2
   292: 'Carrier 04 Duplicate Carrier Number Fault', class No Acknowledgement, trigger "DB302_HMI_Faults_Carrier4_Faults_2" bit 3
   293: 'Spare_Fault_293', class No Acknowledgement, trigger "DB302_HMI_Faults_Carrier4_Faults_2" bit 4
   294: 'Spare_Fault_294', class No Acknowledgement, trigger "DB302_HMI_Faults_Carrier4_Faults_2" bit 5
   295: 'Spare_Fault_295', class No Acknowledgement, trigger "DB302_HMI_Faults_Carrier4_Faults_2" bit 6
   296: 'Spare_Fault_296', class No Acknowledgement, trigger "DB302_HMI_Faults_Carrier4_Faults_2" bit 7
   297: 'Spare_Fault_297', class No Acknowledgement, trigger "DB302_HMI_Faults_Carrier4_Faults_2" bit 8
   298: 'Spare_Fault_298', class No Acknowledgement, trigger "DB302_HMI_Faults_Carrier4_Faults_2" bit 9
   299: 'Spare_Fault_299', class No Acknowledgement, trigger "DB302_HMI_Faults_Carrier4_Faults_2" bit 10
   300: 'Spare_Fault_300', class No Acknowledgement, trigger "DB302_HMI_Faults_Carrier4_Faults_2" bit 11
   301: 'Spare_Fault_301', class No Acknowledgement, trigger "DB302_HMI_Faults_Carrier4_Faults_2" bit 12
   302: 'Spare_Fault_302', class No Acknowledgement, trigger "DB302_HMI_Faults_Carrier4_Faults_2" bit 13
   303: 'Spare_Fault_303', class No Acknowledgement, trigger "DB302_HMI_Faults_Carrier4_Faults_2" bit 14
   304: 'Spare_Fault_304', class No Acknowledgement, trigger "DB302_HMI_Faults_Carrier4_Faults_2" bit 15
   305: 'Spare_Fault_305', class No Acknowledgement, trigger "DB302_HMI_Faults_Carrier4_Faults_3" bit 0
   306: 'Spare_Fault_306', class No Acknowledgement, trigger "DB302_HMI_Faults_Carrier4_Faults_3" bit 1
   307: 'Spare_Fault_307', class No Acknowledgement, trigger "DB302_HMI_Faults_Carrier4_Faults_3" bit 2
   308: 'Spare_Fault_308', class No Acknowledgement, trigger "DB302_HMI_Faults_Carrier4_Faults_3" bit 3
   309: 'Spare_Fault_309', class No Acknowledgement, trigger "DB302_HMI_Faults_Carrier4_Faults_3" bit 4
   310: 'Spare_Fault_310', class No Acknowledgement, trigger "DB302_HMI_Faults_Carrier4_Faults_3" bit 5
   311: 'Spare_Fault_311', class No Acknowledgement, trigger "DB302_HMI_Faults_Carrier4_Faults_3" bit 6
   312: 'Spare_Fault_312', class No Acknowledgement, trigger "DB302_HMI_Faults_Carrier4_Faults_3" bit 7
   313: 'Spare_Fault_313', class No Acknowledgement, trigger "DB302_HMI_Faults_Carrier4_Faults_3" bit 8
   314: 'Spare_Fault_314', class No Acknowledgement, trigger "DB302_HMI_Faults_Carrier4_Faults_3" bit 9
   315: 'Spare_Fault_315', class No Acknowledgement, trigger "DB302_HMI_Faults_Carrier4_Faults_3" bit 10
   316: 'Spare_Fault_316', class No Acknowledgement, trigger "DB302_HMI_Faults_Carrier4_Faults_3" bit 11
   317: 'Spare_Fault_317', class No Acknowledgement, trigger "DB302_HMI_Faults_Carrier4_Faults_3" bit 12
   318: 'Spare_Fault_318', class No Acknowledgement, trigger "DB302_HMI_Faults_Carrier4_Faults_3" bit 13
   319: 'Spare_Fault_319', class No Acknowledgement, trigger "DB302_HMI_Faults_Carrier4_Faults_3" bit 14
   320: 'Spare_Fault_320', class No Acknowledgement, trigger "DB302_HMI_Faults_Carrier4_Faults_3" bit 15
   321: 'Carrier 05 Disconnect Open Power Fault DI11.0', class No Acknowledgement, trigger "DB302_HMI_Faults_Carrier5_Faults_0" bit 0
   322: 'Carrier 05 Drive Profinet Comm Fault', class No Acknowledgement, trigger "DB302_HMI_Faults_Carrier5_Faults_0" bit 1
   323: 'Carrier 05 Production Stop Not Reset', class No Acknowledgement, trigger "DB302_HMI_Faults_Carrier5_Faults_0" bit 2
   324: 'Carrier 05 CB02122 Tripped', class No Acknowledgement, trigger "DB302_HMI_Faults_Carrier5_Faults_0" bit 3
   325: 'Carrier 05 CB02123 Tripped', class No Acknowledgement, trigger "DB302_HMI_Faults_Carrier5_Faults_0" bit 4
   326: 'Carrier 05 AUX1 CB Tripped', class No Acknowledgement, trigger "DB302_HMI_Faults_Carrier5_Faults_0" bit 5
   327: 'Carrier 05 AUX2 CB Tripped', class No Acknowledgement, trigger "DB302_HMI_Faults_Carrier5_Faults_0" bit 6
   328: 'Carrier 05 PLC Not Communicating', class No Acknowledgement, trigger "DB302_HMI_Faults_Carrier5_Faults_0" bit 7
   329: 'Carrier 05 Safe Input Card Fault', class No Acknowledgement, trigger "DB302_HMI_Faults_Carrier5_Faults_0" bit 8
   330: 'Carrier 05 Safe Output Card Fault', class No Acknowledgement, trigger "DB302_HMI_Faults_Carrier5_Faults_0" bit 9
   331: 'Carrier 05 Standard Input Card Fault', class No Acknowledgement, trigger "DB302_HMI_Faults_Carrier5_Faults_0" bit 10
   332: 'Carrier 05 Standard Output Card Fault', class No Acknowledgement, trigger "DB302_HMI_Faults_Carrier5_Faults_0" bit 11
   333: 'Carrier 05 Encoder Position Fault', class No Acknowledgement, trigger "DB302_HMI_Faults_Carrier5_Faults_0" bit 12
   334: 'Carrier 05 Encoder Internal Error', class No Acknowledgement, trigger "DB302_HMI_Faults_Carrier5_Faults_0" bit 13
   335: 'Carrier 05 Encoder Comm Fault', class No Acknowledgement, trigger "DB302_HMI_Faults_Carrier5_Faults_0" bit 14
   336: 'Carrier 05 HMI Comm Fault', class No Acknowledgement, trigger "DB302_HMI_Faults_Carrier5_Faults_0" bit 15
   337: 'Carrier 05 Crash Detection Fault', class No Acknowledgement, trigger "DB302_HMI_Faults_Carrier5_Faults_1" bit 0
   338: 'Carrier 05 Carrier Number Invalid', class No Acknowledgement, trigger "DB302_HMI_Faults_Carrier5_Faults_1" bit 1
   339: 'Carrier 05 Drive: PROFINET configuration error', class No Acknowledgement, trigger "DB302_HMI_Faults_Carrier5_Faults_1" bit 2
   340: 'Carrier 05 Drive: Error internal communications', class No Acknowledgement, trigger "DB302_HMI_Faults_Carrier5_Faults_1" bit 3
   341: 'Carrier 05 Drive: Motor overtemperature', class No Acknowledgement, trigger "DB302_HMI_Faults_Carrier5_Faults_1" bit 4
   342: 'Carrier 05 Drive: Motor overcurrent', class No Acknowledgement, trigger "DB302_HMI_Faults_Carrier5_Faults_1" bit 5
   343: 'Carrier 05 Drive: Infeed or power unit not ready', class No Acknowledgement, trigger "DB302_HMI_Faults_Carrier5_Faults_1" bit 6
   344: 'Carrier 05 Drive: Short-circuit/ground fault detected', class No Acknowledgement, trigger "DB302_HMI_Faults_Carrier5_Faults_1" bit 7
   345: 'Carrier 05 Drive: PROFINET Setpoint timeout', class No Acknowledgement, trigger "DB302_HMI_Faults_Carrier5_Faults_1" bit 8
   346: 'Carrier 05 Power unit: Overcurrent', class No Acknowledgement, trigger "DB302_HMI_Faults_Carrier5_Faults_1" bit 9
   347: 'Carrier 05 Power unit: DC link voltage overvoltage', class No Acknowledgement, trigger "DB302_HMI_Faults_Carrier5_Faults_1" bit 10
   348: 'Carrier 05 Power unit: DC link voltage undervoltage', class No Acknowledgement, trigger "DB302_HMI_Faults_Carrier5_Faults_1" bit 11
   349: 'Carrier 05 Power unit: Line phase failure in main circuit', class No Acknowledgement, trigger "DB302_HMI_Faults_Carrier5_Faults_1" bit 12
   350: 'Carrier 05 Power unit: Phase failure motor cable', class No Acknowledgement, trigger "DB302_HMI_Faults_Carrier5_Faults_1" bit 13
   351: 'Carrier 05 Power unit: Ground fault', class No Acknowledgement, trigger "DB302_HMI_Faults_Carrier5_Faults_1" bit 14
   352: 'Spare_Fault_352', class No Acknowledgement, trigger "DB302_HMI_Faults_Carrier5_Faults_1" bit 15
   353: 'Carrier 05 Motion Off Fault', class No Acknowledgement, trigger "DB302_HMI_Faults_Carrier5_Faults_2" bit 0
   354: 'Carrier 05 Motion On Fault', class No Acknowledgement, trigger "DB302_HMI_Faults_Carrier5_Faults_2" bit 1
   355: 'Carrier 05 Spacing Fault', class No Acknowledgement, trigger "DB302_HMI_Faults_Carrier5_Faults_2" bit 2
   356: 'Carrier 05 Duplicate Carrier Number Fault', class No Acknowledgement, trigger "DB302_HMI_Faults_Carrier5_Faults_2" bit 3
   357: 'Spare_Fault_357', class No Acknowledgement, trigger "DB302_HMI_Faults_Carrier5_Faults_2" bit 4
   358: 'Spare_Fault_358', class No Acknowledgement, trigger "DB302_HMI_Faults_Carrier5_Faults_2" bit 5
   359: 'Spare_Fault_359', class No Acknowledgement, trigger "DB302_HMI_Faults_Carrier5_Faults_2" bit 6
   360: 'Spare_Fault_360', class No Acknowledgement, trigger "DB302_HMI_Faults_Carrier5_Faults_2" bit 7
   361: 'Spare_Fault_361', class No Acknowledgement, trigger "DB302_HMI_Faults_Carrier5_Faults_2" bit 8
   362: 'Spare_Fault_362', class No Acknowledgement, trigger "DB302_HMI_Faults_Carrier5_Faults_2" bit 9
   363: 'Spare_Fault_363', class No Acknowledgement, trigger "DB302_HMI_Faults_Carrier5_Faults_2" bit 10
   364: 'Spare_Fault_364', class No Acknowledgement, trigger "DB302_HMI_Faults_Carrier5_Faults_2" bit 11
   365: 'Spare_Fault_365', class No Acknowledgement, trigger "DB302_HMI_Faults_Carrier5_Faults_2" bit 12
   366: 'Spare_Fault_366', class No Acknowledgement, trigger "DB302_HMI_Faults_Carrier5_Faults_2" bit 13
   367: 'Spare_Fault_367', class No Acknowledgement, trigger "DB302_HMI_Faults_Carrier5_Faults_2" bit 14
   368: 'Spare_Fault_368', class No Acknowledgement, trigger "DB302_HMI_Faults_Carrier5_Faults_2" bit 15
   369: 'Spare_Fault_369', class No Acknowledgement, trigger "DB302_HMI_Faults_Carrier5_Faults_3" bit 0
   370: 'Spare_Fault_370', class No Acknowledgement, trigger "DB302_HMI_Faults_Carrier5_Faults_3" bit 1
   371: 'Spare_Fault_371', class No Acknowledgement, trigger "DB302_HMI_Faults_Carrier5_Faults_3" bit 2
   372: 'Spare_Fault_372', class No Acknowledgement, trigger "DB302_HMI_Faults_Carrier5_Faults_3" bit 3
   373: 'Spare_Fault_373', class No Acknowledgement, trigger "DB302_HMI_Faults_Carrier5_Faults_3" bit 4
   374: 'Spare_Fault_374', class No Acknowledgement, trigger "DB302_HMI_Faults_Carrier5_Faults_3" bit 5
   375: 'Spare_Fault_375', class No Acknowledgement, trigger "DB302_HMI_Faults_Carrier5_Faults_3" bit 6
   376: 'Spare_Fault_376', class No Acknowledgement, trigger "DB302_HMI_Faults_Carrier5_Faults_3" bit 7
   377: 'Spare_Fault_377', class No Acknowledgement, trigger "DB302_HMI_Faults_Carrier5_Faults_3" bit 8
   378: 'Spare_Fault_378', class No Acknowledgement, trigger "DB302_HMI_Faults_Carrier5_Faults_3" bit 9
   379: 'Spare_Fault_379', class No Acknowledgement, trigger "DB302_HMI_Faults_Carrier5_Faults_3" bit 10
   380: 'Spare_Fault_380', class No Acknowledgement, trigger "DB302_HMI_Faults_Carrier5_Faults_3" bit 11
   381: 'Spare_Fault_381', class No Acknowledgement, trigger "DB302_HMI_Faults_Carrier5_Faults_3" bit 12
   382: 'Spare_Fault_382', class No Acknowledgement, trigger "DB302_HMI_Faults_Carrier5_Faults_3" bit 13
   383: 'Spare_Fault_383', class No Acknowledgement, trigger "DB302_HMI_Faults_Carrier5_Faults_3" bit 14
   384: 'Spare_Fault_384', class No Acknowledgement, trigger "DB302_HMI_Faults_Carrier5_Faults_3" bit 15
   385: 'Carrier 06 Disconnect Open Power Fault DI11.0', class No Acknowledgement, trigger "DB302_HMI_Faults_Carrier6_Faults_0" bit 0
   386: 'Carrier 06 Drive Profinet Comm Fault', class No Acknowledgement, trigger "DB302_HMI_Faults_Carrier6_Faults_0" bit 1
   387: 'Carrier 06 Production Stop Not Reset', class No Acknowledgement, trigger "DB302_HMI_Faults_Carrier6_Faults_0" bit 2
   388: 'Carrier 06 CB02122 Tripped', class No Acknowledgement, trigger "DB302_HMI_Faults_Carrier6_Faults_0" bit 3
   389: 'Carrier 06 CB02123 Tripped', class No Acknowledgement, trigger "DB302_HMI_Faults_Carrier6_Faults_0" bit 4
   390: 'Carrier 06 AUX1 CB Tripped', class No Acknowledgement, trigger "DB302_HMI_Faults_Carrier6_Faults_0" bit 5
   391: 'Carrier 06 AUX2 CB Tripped', class No Acknowledgement, trigger "DB302_HMI_Faults_Carrier6_Faults_0" bit 6
   392: 'Carrier 06 PLC Not Communicating', class No Acknowledgement, trigger "DB302_HMI_Faults_Carrier6_Faults_0" bit 7
   393: 'Carrier 06 Safe Input Card Fault', class No Acknowledgement, trigger "DB302_HMI_Faults_Carrier6_Faults_0" bit 8
   394: 'Carrier 06 Safe Output Card Fault', class No Acknowledgement, trigger "DB302_HMI_Faults_Carrier6_Faults_0" bit 9
   395: 'Carrier 06 Standard Input Card Fault', class No Acknowledgement, trigger "DB302_HMI_Faults_Carrier6_Faults_0" bit 10
   396: 'Carrier 06 Standard Output Card Fault', class No Acknowledgement, trigger "DB302_HMI_Faults_Carrier6_Faults_0" bit 11
   397: 'Carrier 06 Encoder Position Fault', class No Acknowledgement, trigger "DB302_HMI_Faults_Carrier6_Faults_0" bit 12
   398: 'Carrier 06 Encoder Internal Error', class No Acknowledgement, trigger "DB302_HMI_Faults_Carrier6_Faults_0" bit 13
   399: 'Carrier 06 Encoder Comm Fault', class No Acknowledgement, trigger "DB302_HMI_Faults_Carrier6_Faults_0" bit 14
   400: 'Carrier 06 HMI Comm Fault', class No Acknowledgement, trigger "DB302_HMI_Faults_Carrier6_Faults_0" bit 15
   401: 'Carrier 06 Crash Detection Fault', class No Acknowledgement, trigger "DB302_HMI_Faults_Carrier6_Faults_1" bit 0
   402: 'Carrier 06 Carrier Number Invalid', class No Acknowledgement, trigger "DB302_HMI_Faults_Carrier6_Faults_1" bit 1
   403: 'Carrier 06 Drive: PROFINET configuration error', class No Acknowledgement, trigger "DB302_HMI_Faults_Carrier6_Faults_1" bit 2
   404: 'Carrier 06 Drive: Error internal communications', class No Acknowledgement, trigger "DB302_HMI_Faults_Carrier6_Faults_1" bit 3
   405: 'Carrier 06 Drive: Motor overtemperature', class No Acknowledgement, trigger "DB302_HMI_Faults_Carrier6_Faults_1" bit 4
   406: 'Carrier 06 Drive: Motor overcurrent', class No Acknowledgement, trigger "DB302_HMI_Faults_Carrier6_Faults_1" bit 5
   407: 'Carrier 06 Drive: Infeed or power unit not ready', class No Acknowledgement, trigger "DB302_HMI_Faults_Carrier6_Faults_1" bit 6
   408: 'Carrier 06 Drive: Short-circuit/ground fault detected', class No Acknowledgement, trigger "DB302_HMI_Faults_Carrier6_Faults_1" bit 7
   409: 'Carrier 06 Drive: PROFINET Setpoint timeout', class No Acknowledgement, trigger "DB302_HMI_Faults_Carrier6_Faults_1" bit 8
   410: 'Carrier 06 Power unit: Overcurrent', class No Acknowledgement, trigger "DB302_HMI_Faults_Carrier6_Faults_1" bit 9
   411: 'Carrier 06 Power unit: DC link voltage overvoltage', class No Acknowledgement, trigger "DB302_HMI_Faults_Carrier6_Faults_1" bit 10
   412: 'Carrier 06 Power unit: DC link voltage undervoltage', class No Acknowledgement, trigger "DB302_HMI_Faults_Carrier6_Faults_1" bit 11
   413: 'Carrier 06 Power unit: Line phase failure in main circuit', class No Acknowledgement, trigger "DB302_HMI_Faults_Carrier6_Faults_1" bit 12
   414: 'Carrier 06 Power unit: Phase failure motor cable', class No Acknowledgement, trigger "DB302_HMI_Faults_Carrier6_Faults_1" bit 13
   415: 'Carrier 06 Power unit: Ground fault', class No Acknowledgement, trigger "DB302_HMI_Faults_Carrier6_Faults_1" bit 14
   416: 'Spare_Fault_416', class No Acknowledgement, trigger "DB302_HMI_Faults_Carrier6_Faults_1" bit 15
   417: 'Carrier 06 Motion Off Fault', class No Acknowledgement, trigger "DB302_HMI_Faults_Carrier6_Faults_2" bit 0
   418: 'Carrier 06 Motion On Fault', class No Acknowledgement, trigger "DB302_HMI_Faults_Carrier6_Faults_2" bit 1
   419: 'Carrier 06 Spacing Fault', class No Acknowledgement, trigger "DB302_HMI_Faults_Carrier6_Faults_2" bit 2
   420: 'Carrier 06 Duplicate Carrier Number Fault', class No Acknowledgement, trigger "DB302_HMI_Faults_Carrier6_Faults_2" bit 3
   421: 'Spare_Fault_421', class No Acknowledgement, trigger "DB302_HMI_Faults_Carrier6_Faults_2" bit 4
   422: 'Spare_Fault_422', class No Acknowledgement, trigger "DB302_HMI_Faults_Carrier6_Faults_2" bit 5
   423: 'Spare_Fault_423', class No Acknowledgement, trigger "DB302_HMI_Faults_Carrier6_Faults_2" bit 6
   424: 'Spare_Fault_424', class No Acknowledgement, trigger "DB302_HMI_Faults_Carrier6_Faults_2" bit 7
   425: 'Spare_Fault_425', class No Acknowledgement, trigger "DB302_HMI_Faults_Carrier6_Faults_2" bit 8
   426: 'Spare_Fault_426', class No Acknowledgement, trigger "DB302_HMI_Faults_Carrier6_Faults_2" bit 9
   427: 'Spare_Fault_427', class No Acknowledgement, trigger "DB302_HMI_Faults_Carrier6_Faults_2" bit 10
   428: 'Spare_Fault_428', class No Acknowledgement, trigger "DB302_HMI_Faults_Carrier6_Faults_2" bit 11
   429: 'Spare_Fault_429', class No Acknowledgement, trigger "DB302_HMI_Faults_Carrier6_Faults_2" bit 12
   430: 'Spare_Fault_430', class No Acknowledgement, trigger "DB302_HMI_Faults_Carrier6_Faults_2" bit 13
   431: 'Spare_Fault_431', class No Acknowledgement, trigger "DB302_HMI_Faults_Carrier6_Faults_2" bit 14
   432: 'Spare_Fault_432', class No Acknowledgement, trigger "DB302_HMI_Faults_Carrier6_Faults_2" bit 15
   433: 'Spare_Fault_433', class No Acknowledgement, trigger "DB302_HMI_Faults_Carrier6_Faults_3" bit 0
   434: 'Spare_Fault_434', class No Acknowledgement, trigger "DB302_HMI_Faults_Carrier6_Faults_3" bit 1
   435: 'Spare_Fault_435', class No Acknowledgement, trigger "DB302_HMI_Faults_Carrier6_Faults_3" bit 2
   436: 'Spare_Fault_436', class No Acknowledgement, trigger "DB302_HMI_Faults_Carrier6_Faults_3" bit 3
   437: 'Spare_Fault_437', class No Acknowledgement, trigger "DB302_HMI_Faults_Carrier6_Faults_3" bit 4